// TIA Portal project "Ampelanlage_1" (V20)

(* hardware
DEVICE "S7-1500/ET200MP-Station_1"  S7-1500 station
   slot 0: "Profilschiene_0"  Rack  6ES7 590-1***0-0AA0
   slot 1: "PLC_1"  CPU 1513-1 PN  6ES7 513-1AM03-0AB0  V4.0
      slot 3: "CPU-Display_1"  6ES7591-1AA00-0AA0
      slot 32768: "PROFINET-Schnittstelle_1"  X1
         slot 32769: "Port_1"  X1 P1
         slot 32770: "Port_2"  X1 P2
      slot 34817: "Virtual CP interface port_1"  Virtual CP interface port  Virtual CP interface port FW V4.0
   slot 2: "DI 16x24VDC BA_1"  DI 16x24VDC BA  6ES7 521-1BH10-0AA0  V1.1
   slot 3: "DQ 16x24VDC/0.5A ST_1"  DQ 16x24VDC/0.5A ST  6ES7 522-1BH00-0AB0  V2.0
   slot 4: "AI 8xU/I/R/RTD BA_2"  AI 8xU/I/R/RTD BA  6ES7 531-7QF00-0AB0  V1.0
   slot 5: "AQ 8xU/I HS_2"  AQ 8xU/I HS  6ES7 532-5HF00-0AB0  V2.2
DEVICE "HMI_1"  TP700 Comfort
   slot 0: "HMI_1"  TP700 Comfort  6AV2 124-0GC01-0AX0  17.0.0.0
   slot 1: "HMI_RT_1"  TP700 Comfort  6AV2 124-0GC01-0AX0  17.0.0.0
   slot 5: "HMI_1.IE_CP_1"  PROFINET Interface  17.0.0.0
      slot 1: "PROFINET Schnittstelle_1"  PROFINET Interface
         slot 1: "Port_1"  Port
         slot 2: "Port_2"  Port
   slot 7: "HMI_1.MPI/DP_CP_1"  MPI/DP Interface  17.0.0.0
*)

// ===== PLC "PLC_1"  CPU 1513-1 PN =====

VAR_GLOBAL   // PLC tag table "Eingaenge"
   "S1" AT %E0.0 : Bool;   // Starttaster
END_VAR

VAR_GLOBAL   // PLC tag table "Ausgaenge"
   "1H1" AT %A0.0 : Bool;   // Hauptstraße 1 (rot)
   "1H2" AT %A0.1 : Bool;   // Hauptstraße 1 (gelb)
   "1H3" AT %A0.2 : Bool;   // Hauptstraße 1 (grün)
   "2H1" AT %A0.3 : Bool;   // Hauptstraße 2 (rot)
   "2H2" AT %A0.4 : Bool;   // Hauptstraße 2 (gelb)
   "2H3" AT %A0.5 : Bool;   // Hauptstraße 2 (grün)
   "3H1" AT %A0.6 : Bool;   // Nebenstraße 1 (rot)
   "3H2" AT %A0.7 : Bool;   // Nebenstraße 1 (gelb)
   "3H3" AT %A1.0 : Bool;   // Nebenstraße 1 (grün)
   "4H1" AT %A1.1 : Bool;   // Nebenstraße 2 (rot)
   "4H2" AT %A1.2 : Bool;   // Nebenstraße 2 (gelb)
   "4H3" AT %A1.3 : Bool;   // Nebenstraße 2 (grün)
   "5H1" AT %A1.4 : Bool;   // Fußgänger 1 (rot)
   "5H2" AT %A1.5 : Bool;   // Fußgänger 1 (grün)
   "6H1" AT %A1.6 : Bool;   // Fußgänger 2 (rot)
   "6H2" AT %A1.7 : Bool;   // Fußgänger 2 (grün)
END_VAR

TYPE "typSignale"
   STRUCT
      Hauptstrasse : Struct
         Rot : Bool;   // Hauptstraße Ampel (rot)
         Gelb : Bool;   // Hauptstraße Ampel (gelb)
         Gruen : Bool;   // Hauptstraße Ampel (grün)
      END_STRUCT;
      Nebenstrasse : Struct
         Rot : Bool;   // Nebenstraße Ampel (rot)
         Gelb : Bool;   // Nebenstraße Ampel (gelb)
         Gruen : Bool;   // Nebenstraße Ampel (grün)
      END_STRUCT;
      Fussgaenger : Struct
         Rot : Bool;   // Fußgänger Ampel (rot)
         Gruen : Bool;   // Fußgänger Ampel (grün)
      END_STRUCT;
   END_STRUCT;
END_TYPE

TYPE "typPhasen"
   STRUCT
      Phase_1 : Struct
         NR : UDInt := 1;
         Phasen_Zeit : Time := T#3s;
         Aktiv : Bool;
      END_STRUCT;
      Phase_2 : Struct
         NR : UDInt := 2;
         Phasen_Zeit : Time := T#2s;
         Aktiv : Bool;
      END_STRUCT;
      Phase_3 : Struct
         NR : UDInt := 3;
         Phasen_Zeit : Time := T#10s;
         Aktiv : Bool;
      END_STRUCT;
      Phase_4 : Struct
         NR : UDInt := 4;
         Phasen_Zeit : Time := T#2s;
         Aktiv : Bool;
      END_STRUCT;
      Phase_5 : Struct
         NR : UDInt := 5;
         Phasen_Zeit : Time := T#3s;
         Aktiv : Bool;
      END_STRUCT;
      Phase_6 : Struct
         NR : UDInt := 6;
         Phasen_Zeit : Time := T#2s;
         Aktiv : Bool;
      END_STRUCT;
      Phase_7 : Struct
         NR : UDInt := 7;
         Phasen_Zeit : Time := T#8s;
         Aktiv : Bool;
      END_STRUCT;
      Phase_8 : Struct
         NR : UDInt := 8;
         Phasen_Zeit : Time := T#2s;
         Aktiv : Bool;
      END_STRUCT;
   END_STRUCT;
END_TYPE

TYPE "typTransitionen"
   STRUCT
      Phasen_Transitionen : Struct
         P_1_2 : Bool;
         P_2_3 : Bool;
         P_3_4 : Bool;
         P_4_5 : Bool;
         P_5_6 : Bool;
         P_6_7 : Bool;
         P_7_8 : Bool;
      END_STRUCT;
      Schritt_Transitionen : Struct
         T_0_1 : Bool;
         T_1_2 : Bool;
         T_2_0 : Bool;
         T_2_1 : Bool;
      END_STRUCT;
   END_STRUCT;
END_TYPE

DATA_BLOCK "HMI_Schnittstelle"   // DB1
{ S7_Optimized_Access := 'TRUE' }
VERSION : 0.1
   VAR
      Eingänge : Struct
         S1 : Bool;   // Schalter S1
      END_STRUCT;
      Ausgänge : Struct
         Signale : "typSignale";
      END_STRUCT;
      Schritt_Nr : DInt;
      Ampelphase : Time;
      Phasen : "typPhasen";
      Transitionen : "typTransitionen";
      Anlage_ein : Bool;
   END_VAR
BEGIN
END_DATA_BLOCK

DATA_BLOCK "IDB_Schritte_Ampelanlage"   // DB2
{ S7_Optimized_Access := 'TRUE' }
VERSION : 0.1
// stored: InstanceOfName Prog_Schrittkette_Ampelanlage
"Prog_Schrittkette_Ampelanlage"
BEGIN
END_DATA_BLOCK

FUNCTION_BLOCK "Prog_Schrittkette_Ampelanlage"   // FB1, FBD
{ S7_Optimized_Access := 'TRUE' }
VERSION : 0.1
   VAR_INPUT
      eStart : Bool;
   END_VAR
   VAR_OUTPUT
      aSchritt_Nr : DInt;
   END_VAR
   VAR_IN_OUT
      eaPhasen : "typPhasen";
      eaTransitionen : "typTransitionen";
      eaPhasenzeit : Array[0..8] of Time;
   END_VAR
   VAR
      Schritt_0 : Bool := true;   // 0: Initialschritt
      Schritt_1 : Bool;   // 1: Ampelphase 1
      Schritt_2 : Bool;   // 8: Ampelphase 8
      TOF_Schritt1 : TON_TIME;
      TON_Phase1 : TON_TIME;
      TON_Phase2 : TON_TIME;
      TON_Phase3 : TON_TIME;
      TON_Phase4 : TON_TIME;
      TON_Phase5 : TON_TIME;
      TON_Phase6 : TON_TIME;
      TON_Phase7 : TON_TIME;
      TON_Phase8 : TON_TIME;
      RTRIG_Start_Taster : R_TRIG;
      MDB_Phase_1 : "Ampelphase";
      MDB_Phase_2 : "Ampelphase";
      MDB_Phase_3 : "Ampelphase";
      MDB_Phase_4 : "Ampelphase";
      MDB_Phase_5 : "Ampelphase";
      MDB_Phase_6 : "Ampelphase";
      MDB_Phase_7 : "Ampelphase";
      MDB_Phase_8 : "Ampelphase";
      Phasen_gestartet : Bool;
   END_VAR
BEGIN

REGION Network 1: Anlage in Grundstellung
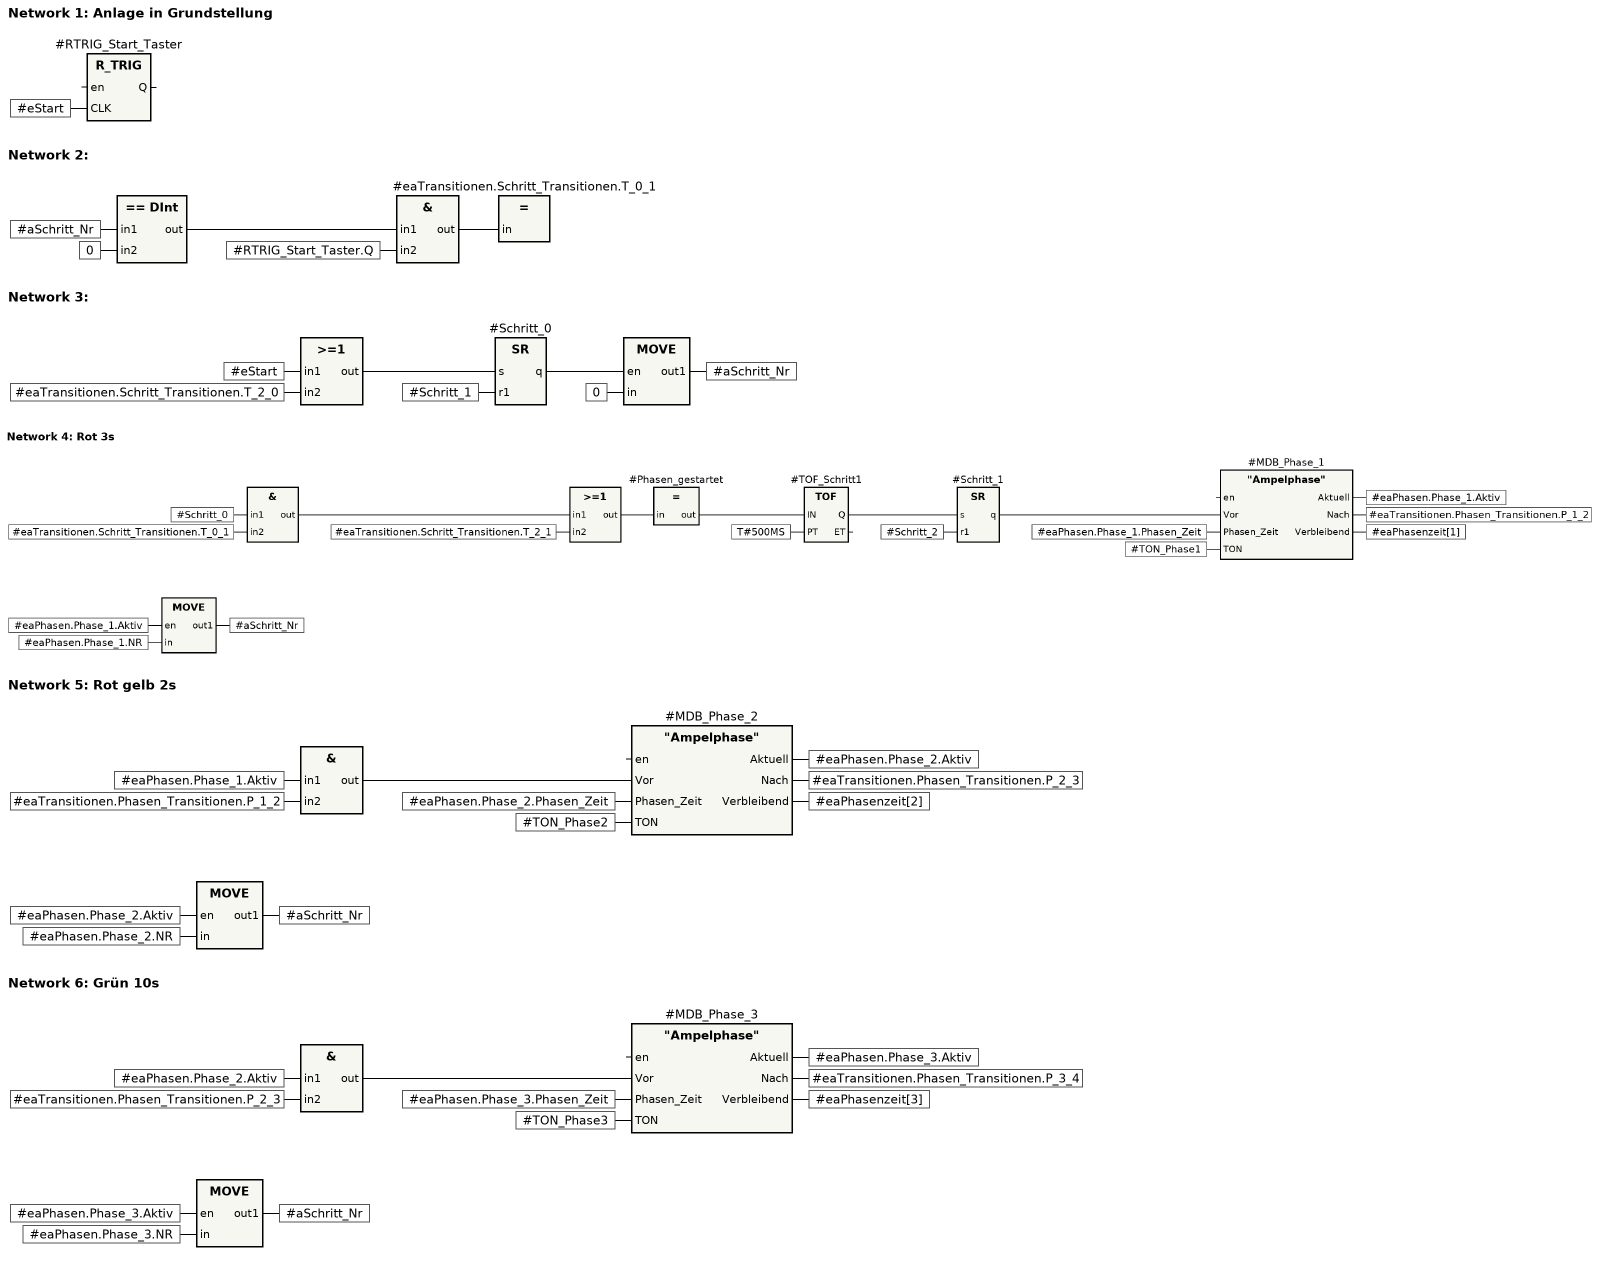
   #RTRIG_Start_Taster(CLK := #eStart);   // R_TRIG
END_REGION

REGION Network 2
   #eaTransitionen.Schritt_Transitionen.T_0_1 := (#aSchritt_Nr = 0) AND #RTRIG_Start_Taster.Q;
END_REGION

REGION Network 3
   IF #eStart OR #eaTransitionen.Schritt_Transitionen.T_2_0 THEN
       #Schritt_0 := TRUE;   // SR flip-flop
   END_IF;
   IF #Schritt_1 THEN #Schritt_0 := FALSE; END_IF;
   IF #Schritt_0 THEN #aSchritt_Nr := 0; END_IF;
END_REGION

REGION Network 4: Rot 3s
   #Phasen_gestartet := (#Schritt_0 AND #eaTransitionen.Schritt_Transitionen.T_0_1) OR #eaTransitionen.Schritt_Transitionen.T_2_1;
   #TOF_Schritt1(IN := #Phasen_gestartet, PT := T#500MS);   // TOF
   IF #TOF_Schritt1.Q THEN
       #Schritt_1 := TRUE;   // SR flip-flop
   END_IF;
   IF #Schritt_2 THEN #Schritt_1 := FALSE; END_IF;
   #MDB_Phase_1(Vor := #Schritt_1,   // "Ampelphase"
                Phasen_Zeit := #eaPhasen.Phase_1.Phasen_Zeit,
                TON := #TON_Phase1,
                Aktuell => #eaPhasen.Phase_1.Aktiv,
                Nach => #eaTransitionen.Phasen_Transitionen.P_1_2,
                Verbleibend => #eaPhasenzeit[1]);
   IF #eaPhasen.Phase_1.Aktiv THEN #aSchritt_Nr := #eaPhasen.Phase_1.NR; END_IF;
END_REGION

REGION Network 5: Rot gelb 2s
   #MDB_Phase_2(Vor := #eaPhasen.Phase_1.Aktiv AND #eaTransitionen.Phasen_Transitionen.P_1_2,   // "Ampelphase"
                Phasen_Zeit := #eaPhasen.Phase_2.Phasen_Zeit,
                TON := #TON_Phase2,
                Aktuell => #eaPhasen.Phase_2.Aktiv,
                Nach => #eaTransitionen.Phasen_Transitionen.P_2_3,
                Verbleibend => #eaPhasenzeit[2]);
   IF #eaPhasen.Phase_2.Aktiv THEN #aSchritt_Nr := #eaPhasen.Phase_2.NR; END_IF;
END_REGION

REGION Network 6: Grün 10s
   #MDB_Phase_3(Vor := #eaPhasen.Phase_2.Aktiv AND #eaTransitionen.Phasen_Transitionen.P_2_3,   // "Ampelphase"
                Phasen_Zeit := #eaPhasen.Phase_3.Phasen_Zeit,
                TON := #TON_Phase3,
                Aktuell => #eaPhasen.Phase_3.Aktiv,
                Nach => #eaTransitionen.Phasen_Transitionen.P_3_4,
                Verbleibend => #eaPhasenzeit[3]);
   IF #eaPhasen.Phase_3.Aktiv THEN #aSchritt_Nr := #eaPhasen.Phase_3.NR; END_IF;
END_REGION

REGION Network 7: Gelb 2s
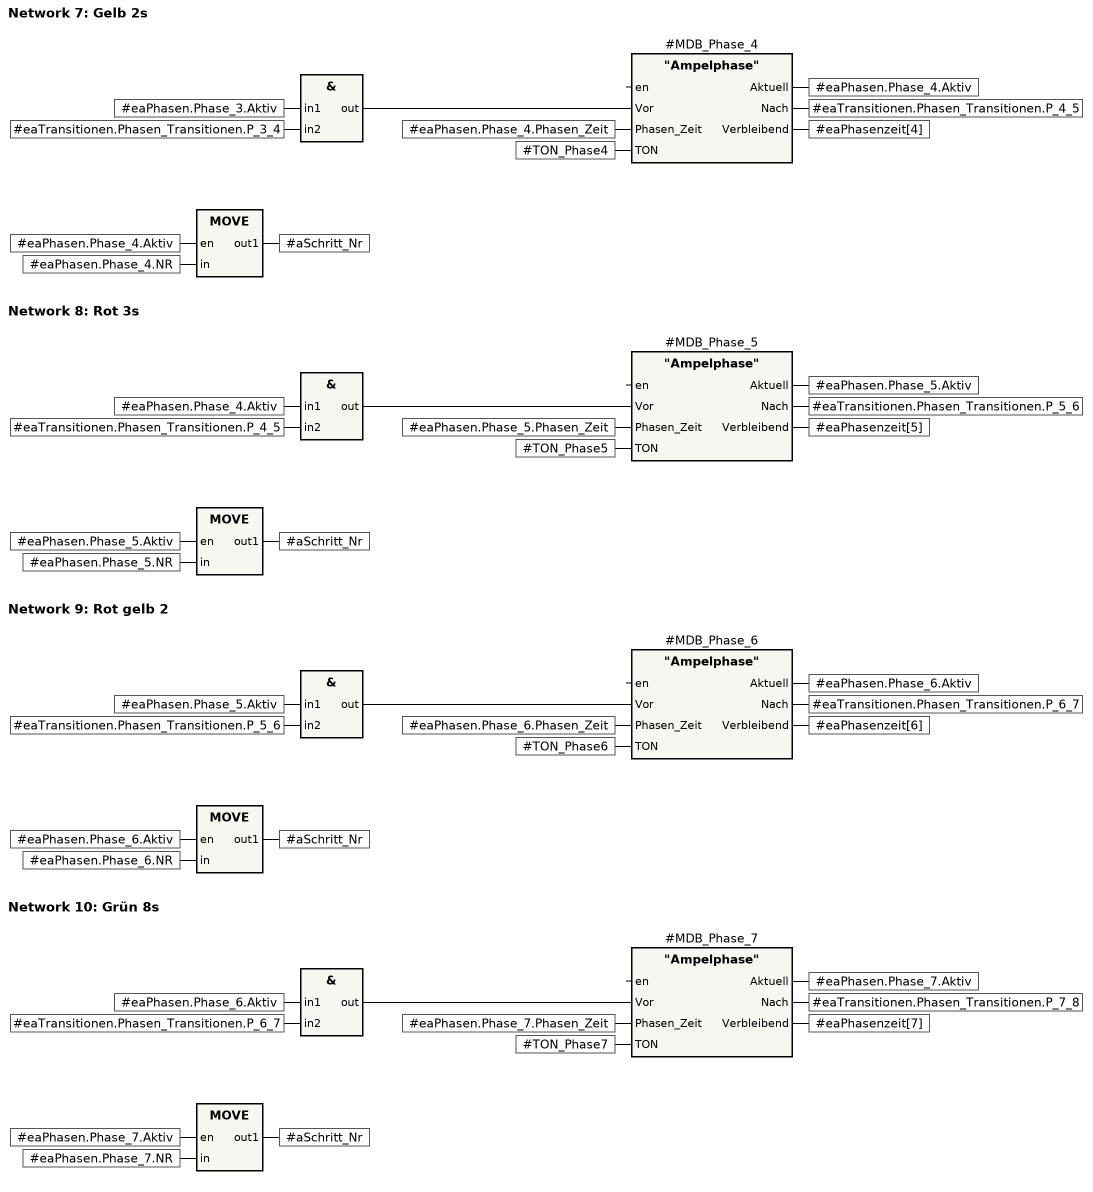
   #MDB_Phase_4(Vor := #eaPhasen.Phase_3.Aktiv AND #eaTransitionen.Phasen_Transitionen.P_3_4,   // "Ampelphase"
                Phasen_Zeit := #eaPhasen.Phase_4.Phasen_Zeit,
                TON := #TON_Phase4,
                Aktuell => #eaPhasen.Phase_4.Aktiv,
                Nach => #eaTransitionen.Phasen_Transitionen.P_4_5,
                Verbleibend => #eaPhasenzeit[4]);
   IF #eaPhasen.Phase_4.Aktiv THEN #aSchritt_Nr := #eaPhasen.Phase_4.NR; END_IF;
END_REGION

REGION Network 8: Rot 3s
   #MDB_Phase_5(Vor := #eaPhasen.Phase_4.Aktiv AND #eaTransitionen.Phasen_Transitionen.P_4_5,   // "Ampelphase"
                Phasen_Zeit := #eaPhasen.Phase_5.Phasen_Zeit,
                TON := #TON_Phase5,
                Aktuell => #eaPhasen.Phase_5.Aktiv,
                Nach => #eaTransitionen.Phasen_Transitionen.P_5_6,
                Verbleibend => #eaPhasenzeit[5]);
   IF #eaPhasen.Phase_5.Aktiv THEN #aSchritt_Nr := #eaPhasen.Phase_5.NR; END_IF;
END_REGION

REGION Network 9: Rot gelb 2
   #MDB_Phase_6(Vor := #eaPhasen.Phase_5.Aktiv AND #eaTransitionen.Phasen_Transitionen.P_5_6,   // "Ampelphase"
                Phasen_Zeit := #eaPhasen.Phase_6.Phasen_Zeit,
                TON := #TON_Phase6,
                Aktuell => #eaPhasen.Phase_6.Aktiv,
                Nach => #eaTransitionen.Phasen_Transitionen.P_6_7,
                Verbleibend => #eaPhasenzeit[6]);
   IF #eaPhasen.Phase_6.Aktiv THEN #aSchritt_Nr := #eaPhasen.Phase_6.NR; END_IF;
END_REGION

REGION Network 10: Grün 8s
   #MDB_Phase_7(Vor := #eaPhasen.Phase_6.Aktiv AND #eaTransitionen.Phasen_Transitionen.P_6_7,   // "Ampelphase"
                Phasen_Zeit := #eaPhasen.Phase_7.Phasen_Zeit,
                TON := #TON_Phase7,
                Aktuell => #eaPhasen.Phase_7.Aktiv,
                Nach => #eaTransitionen.Phasen_Transitionen.P_7_8,
                Verbleibend => #eaPhasenzeit[7]);
   IF #eaPhasen.Phase_7.Aktiv THEN #aSchritt_Nr := #eaPhasen.Phase_7.NR; END_IF;
END_REGION

REGION Network 11: Gelb 2s
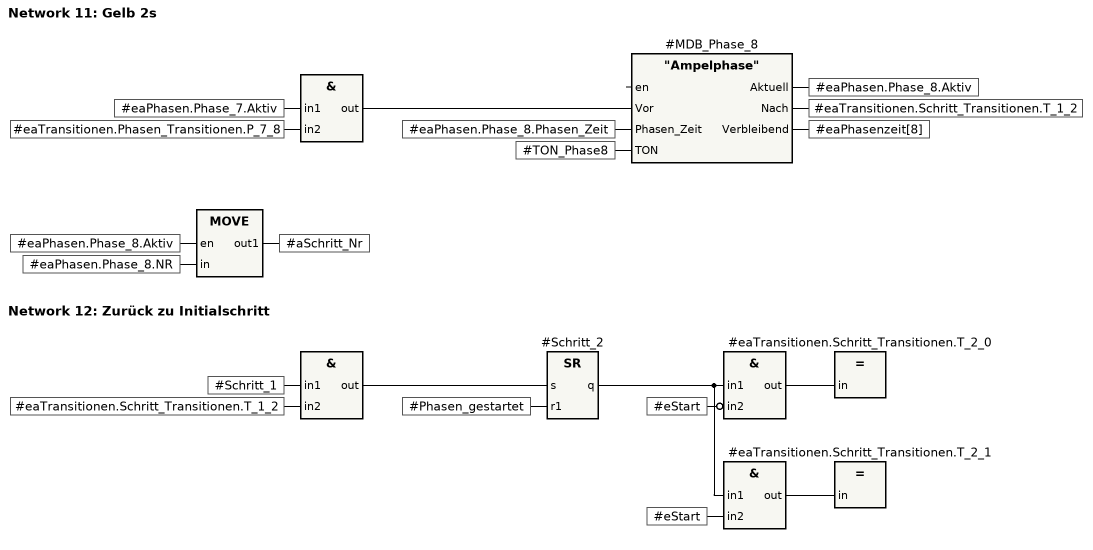
   #MDB_Phase_8(Vor := #eaPhasen.Phase_7.Aktiv AND #eaTransitionen.Phasen_Transitionen.P_7_8,   // "Ampelphase"
                Phasen_Zeit := #eaPhasen.Phase_8.Phasen_Zeit,
                TON := #TON_Phase8,
                Aktuell => #eaPhasen.Phase_8.Aktiv,
                Nach => #eaTransitionen.Schritt_Transitionen.T_1_2,
                Verbleibend => #eaPhasenzeit[8]);
   IF #eaPhasen.Phase_8.Aktiv THEN #aSchritt_Nr := #eaPhasen.Phase_8.NR; END_IF;
END_REGION

REGION Network 12: Zurück zu Initialschritt
   IF #Schritt_1 AND #eaTransitionen.Schritt_Transitionen.T_1_2 THEN
       #Schritt_2 := TRUE;   // SR flip-flop
   END_IF;
   IF #Phasen_gestartet THEN #Schritt_2 := FALSE; END_IF;
   #eaTransitionen.Schritt_Transitionen.T_2_0 := #Schritt_2 AND NOT #eStart;
   #eaTransitionen.Schritt_Transitionen.T_2_1 := #Schritt_2 AND #eStart;
END_REGION
END_FUNCTION_BLOCK

FUNCTION_BLOCK "Ampelphase"   // FB2, FBD
{ S7_Optimized_Access := 'TRUE' }
VERSION : 0.1
   VAR_INPUT
      Vor : Bool;
      Phasen_Zeit : Time;
   END_VAR
   VAR_OUTPUT
      Aktuell : Bool;
      Nach : Bool;
      Verbleibend : Time;
   END_VAR
   VAR_IN_OUT
      TON : TON_TIME;
   END_VAR
BEGIN

REGION Network 1
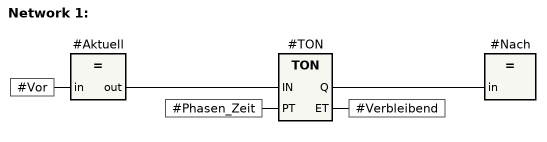
   #Aktuell := #Vor;
   #TON(IN := #Vor, PT := #Phasen_Zeit, ET => #Verbleibend);   // TON
   #Nach := #TON.Q;
END_REGION
END_FUNCTION_BLOCK

FUNCTION_BLOCK "Anlagensignale_einlesen"   // FB3, FBD
{ S7_Optimized_Access := 'TRUE' }
VERSION : 0.1
   VAR
      RTRIG_HMI_Taster : R_TRIG;
      RTRIG_eStart : R_TRIG;
   END_VAR
BEGIN

REGION Network 1: Flankenabfragen
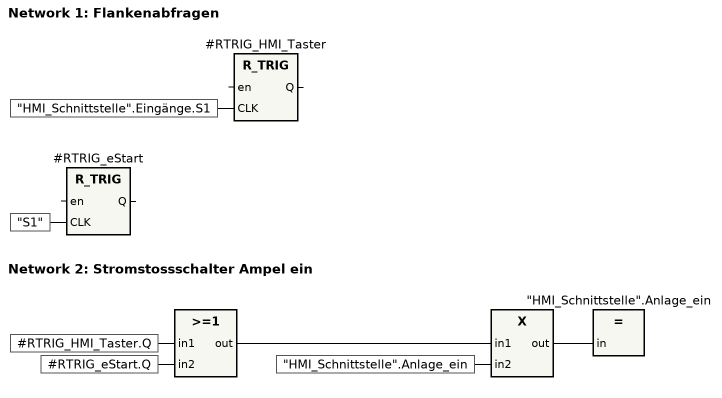
   #RTRIG_HMI_Taster(CLK := "HMI_Schnittstelle".Eingänge.S1);   // R_TRIG
   #RTRIG_eStart(CLK := "S1");   // R_TRIG
END_REGION

REGION Network 2: Stromstossschalter Ampel ein
   "HMI_Schnittstelle".Anlage_ein := (#RTRIG_HMI_Taster.Q OR #RTRIG_eStart.Q) XOR "HMI_Schnittstelle".Anlage_ein;
END_REGION
END_FUNCTION_BLOCK

FUNCTION_BLOCK "Takt"   // FB10101, FBD
TITLE = Taktbaustein parametrierbar
{ S7_Optimized_Access := 'TRUE' }
VERSION : 0.1
// ACHTUNG: keine Zeit darf 0ms sein, ansonsten funktioniert der Baustein nicht.
   VAR_INPUT
      ePulsZeit : Time := T#500MS;   // So lange ist Ausgang = TRUE
      ePauseZeit : Time := T#500MS;   // So lange ist Ausgang = FALSE
   END_VAR
   VAR_OUTPUT
      Q : Bool;
   END_VAR
   VAR
      TP_Puls : TP_TIME;
      TP_Pause : TP_TIME;
   END_VAR
BEGIN

REGION Network 1: Puls Timer
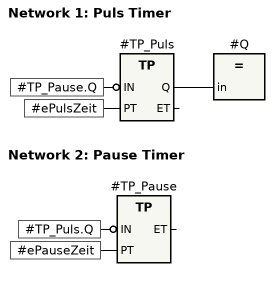
   #TP_Puls(IN := NOT #TP_Pause.Q, PT := #ePulsZeit);   // TP
   #Q := #TP_Puls.Q;
END_REGION

REGION Network 2: Pause Timer
   #TP_Pause(IN := NOT #TP_Puls.Q, PT := #ePauseZeit);   // TP
END_REGION
END_FUNCTION_BLOCK

FUNCTION "Aus_an_Anlage" : Void   // FC1, FBD
{ S7_Optimized_Access := 'TRUE' }
VERSION : 0.1
   VAR_INPUT
      eSignale : "typSignale";
   END_VAR
BEGIN

REGION Network 1: Ampeln Hauptstraße
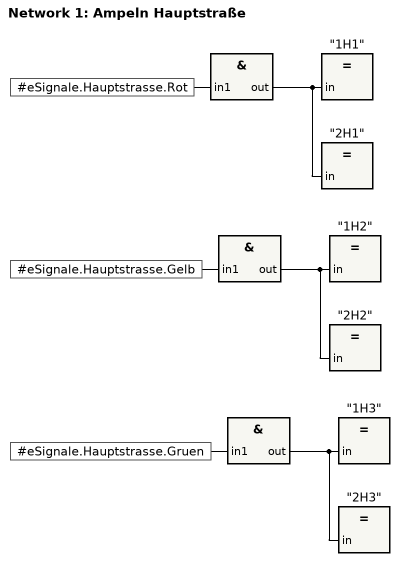
   "1H1" := #eSignale.Hauptstrasse.Rot;
   "2H1" := #eSignale.Hauptstrasse.Rot;
   "1H2" := #eSignale.Hauptstrasse.Gelb;
   "2H2" := #eSignale.Hauptstrasse.Gelb;
   "1H3" := #eSignale.Hauptstrasse.Gruen;
   "2H3" := #eSignale.Hauptstrasse.Gruen;
END_REGION

REGION Network 2 (SCL): Nebenstraße 1 (rot)
   // Ampel Nebenstraße

   "3H1" := "4H1" := #eSignale.Nebenstrasse.Rot;
   "3H2" := "4H2" := #eSignale.Nebenstrasse.Gelb;
   "3H3" := "4H3" := #eSignale.Nebenstrasse.Gruen;


   // Ampel Fussgaenger
   "5H1" := "6H1" := #eSignale.Fussgaenger.Rot;
   "5H2" := "6H2" := #eSignale.Fussgaenger.Gruen;
END_REGION
END_FUNCTION

FUNCTION "Aus_Ampelanlage" : Void   // FC2, FBD
{ S7_Optimized_Access := 'TRUE' }
VERSION : 0.1
   VAR_INPUT
      eSchritt_Nr : DInt;
   END_VAR
   VAR_OUTPUT
      aSignale : "typSignale";
   END_VAR
   VAR_TEMP
      Initialschritt : Bool;
   END_VAR
BEGIN

REGION Network 1
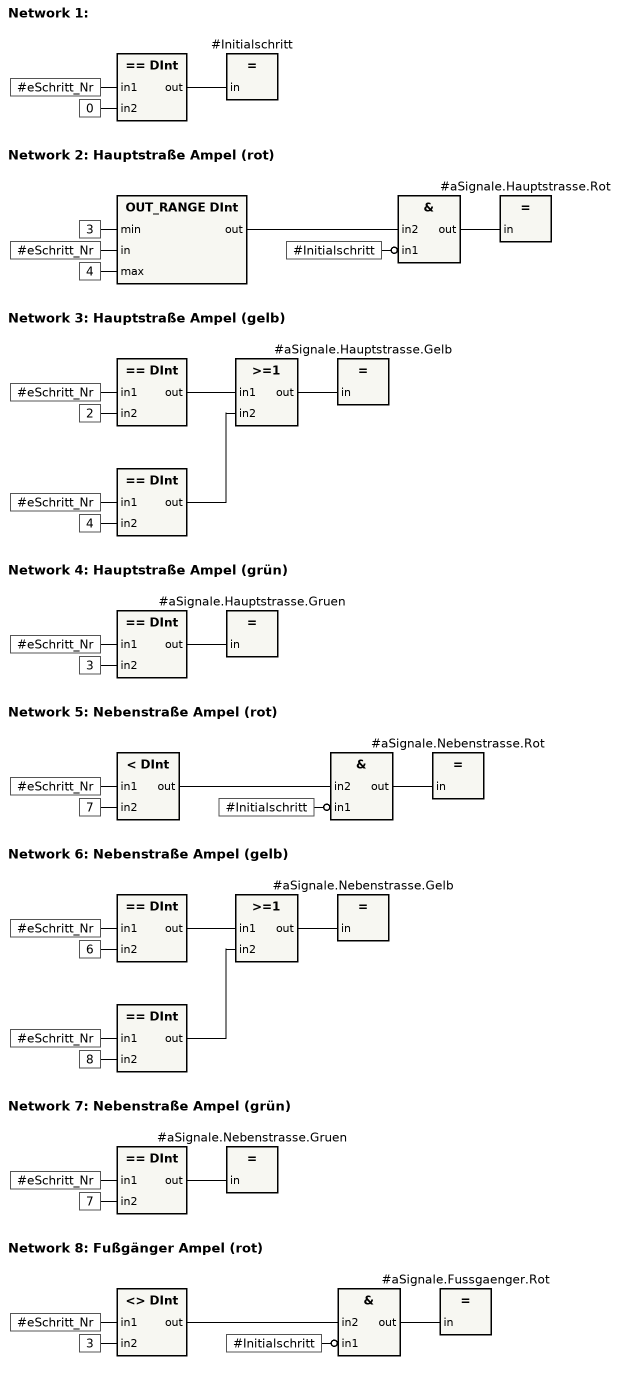
   #Initialschritt := #eSchritt_Nr = 0;
END_REGION

REGION Network 2: Hauptstraße Ampel (rot)
   #aSignale.Hauptstrasse.Rot := ((#eSchritt_Nr < 3) OR (#eSchritt_Nr > 4)) AND NOT #Initialschritt;
END_REGION

REGION Network 3: Hauptstraße Ampel (gelb)
   #aSignale.Hauptstrasse.Gelb := (#eSchritt_Nr = 2) OR (#eSchritt_Nr = 4);
END_REGION

REGION Network 4: Hauptstraße Ampel (grün)
   #aSignale.Hauptstrasse.Gruen := #eSchritt_Nr = 3;
END_REGION

REGION Network 5: Nebenstraße Ampel (rot)
   #aSignale.Nebenstrasse.Rot := (#eSchritt_Nr < 7) AND NOT #Initialschritt;
END_REGION

REGION Network 6: Nebenstraße Ampel (gelb)
   #aSignale.Nebenstrasse.Gelb := (#eSchritt_Nr = 6) OR (#eSchritt_Nr = 8);
END_REGION

REGION Network 7: Nebenstraße Ampel (grün)
   #aSignale.Nebenstrasse.Gruen := #eSchritt_Nr = 7;
END_REGION

REGION Network 8: Fußgänger Ampel (rot)
   #aSignale.Fussgaenger.Rot := (#eSchritt_Nr <> 3) AND NOT #Initialschritt;
END_REGION

REGION Network 9: Fußgänger Ampel (grün)
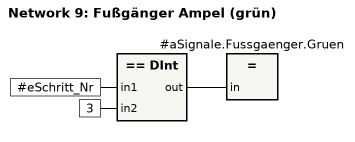
   #aSignale.Fussgaenger.Gruen := #eSchritt_Nr = 3;
END_REGION
END_FUNCTION

ORGANIZATION_BLOCK "Main"   // OB1, FBD, ProgramCycle
TITLE = "Main Program Sweep (Cycle)"
{ S7_Optimized_Access := 'TRUE' }
VERSION : 0.1
   VAR_INPUT
      Initial_Call : Bool;   // Initial call of this OB
      Remanence : Bool;   // =True, if remanent data are available
   END_VAR
   VAR_TEMP
      Phasenzeit : Array[0..8] of Time;
   END_VAR
BEGIN

REGION Network 1
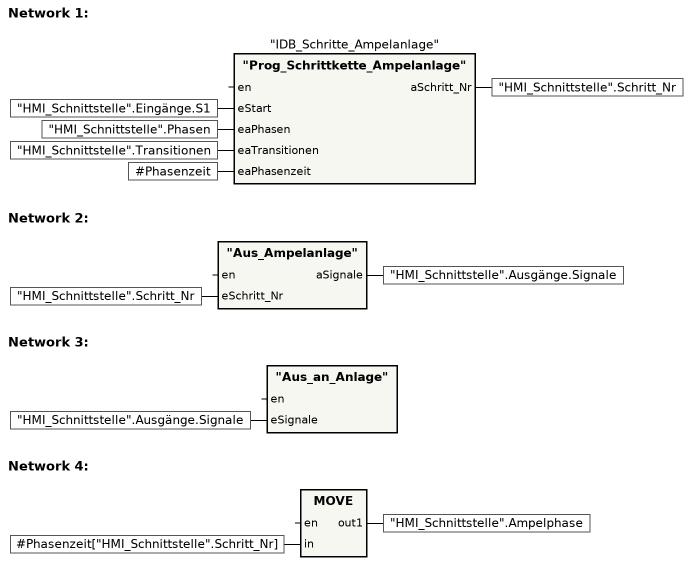
   "IDB_Schritte_Ampelanlage"(eStart := "HMI_Schnittstelle".Eingänge.S1,   // "Prog_Schrittkette_Ampelanlage"
                           eaPhasen := "HMI_Schnittstelle".Phasen,
                           eaTransitionen := "HMI_Schnittstelle".Transitionen,
                           eaPhasenzeit := #Phasenzeit,
                           aSchritt_Nr => "HMI_Schnittstelle".Schritt_Nr);
END_REGION

REGION Network 2
   "Aus_Ampelanlage"(eSchritt_Nr := "HMI_Schnittstelle".Schritt_Nr,
                     aSignale => "HMI_Schnittstelle".Ausgänge.Signale);
END_REGION

REGION Network 3
   "Aus_an_Anlage"(eSignale := "HMI_Schnittstelle".Ausgänge.Signale);
END_REGION

REGION Network 4
   "HMI_Schnittstelle".Ampelphase := #Phasenzeit["HMI_Schnittstelle".Schritt_Nr];
END_REGION
END_ORGANIZATION_BLOCK

(* ===== HMI "HMI_RT_1" =====
system functions are stored by id; their names below are inferred from use
connection "HMI_Verbindung_1": ETHERNET, S7_1500_OMS

HMI tags "Standard-Variablentabelle"
   "HMI_Schnittstelle_S1" : Bool = PLC HMI_Schnittstelle.Eingänge.S1, 500 ms
   "HMI_Schnittstelle_Ausgänge_Schritt_Nr" : DInt = PLC HMI_Schnittstelle.Schritt_Nr, 100 ms
   "HMI_Schnittstelle_Ausgänge_1H1" : Bool = PLC HMI_Schnittstelle.Ausgänge.Signale.Hauptstrasse.Rot, 100 ms
   "HMI_Schnittstelle_Ausgänge_1H2" : Bool = PLC HMI_Schnittstelle.Ausgänge.Signale.Hauptstrasse.Gelb, 100 ms
   "HMI_Schnittstelle_Ausgänge_1H3" : Bool = PLC HMI_Schnittstelle.Ausgänge.Signale.Hauptstrasse.Gruen, 100 ms
   "HMI_Schnittstelle_Ausgänge_2H1" : Bool = PLC HMI_Schnittstelle.Ausgänge.Signale.Nebenstrasse.Rot, 100 ms
   "HMI_Schnittstelle_Ausgänge_2H2" : Bool = PLC HMI_Schnittstelle.Ausgänge.Signale.Nebenstrasse.Gelb, 100 ms
   "HMI_Schnittstelle_Ausgänge_2H3" : Bool = PLC HMI_Schnittstelle.Ausgänge.Signale.Nebenstrasse.Gruen, 100 ms
   "HMI_Schnittstelle_Ausgänge_3H1" : Bool = PLC HMI_Schnittstelle.Ausgänge.Signale.Fussgaenger.Rot, 100 ms
   "HMI_Schnittstelle_Ausgänge_3H2" : Bool = PLC HMI_Schnittstelle.Ausgänge.Signale.Fussgaenger.Gruen, 100 ms
   "HMI_Schnittstelle_Ampelphase" : Time = PLC HMI_Schnittstelle.Ampelphase, 100 ms

screen "Ampelanlage" 800x480
   Button "Schaltfläche_1" at 700,444 size 96x32; TextOff 'S1'
      on Click: InvertBit("HMI_Schnittstelle_S1")
      Appearance <- "HMI_Schnittstelle_S1"
   Circle "Kreis_1" at 286,238 size 16x16
      Appearance <- "HMI_Schnittstelle_Ausgänge_1H1"
   Circle "Kreis_2" at 268,238 size 16x16
      Appearance <- "HMI_Schnittstelle_Ausgänge_1H2"
   Circle "Kreis_3" at 250,238 size 16x16
      Appearance <- "HMI_Schnittstelle_Ausgänge_1H3"
   Circle "Kreis_4" at 498,26 size 16x16
      Appearance <- "HMI_Schnittstelle_Ausgänge_1H1"
   Circle "Kreis_5" at 516,26 size 16x16
      Appearance <- "HMI_Schnittstelle_Ausgänge_1H2"
   Circle "Kreis_6" at 534,26 size 16x16
      Appearance <- "HMI_Schnittstelle_Ausgänge_1H3"
   Circle "Kreis_7" at 498,318 size 16x16
      Appearance <- "HMI_Schnittstelle_Ausgänge_2H1"
   Circle "Kreis_8" at 498,336 size 16x16
      Appearance <- "HMI_Schnittstelle_Ausgänge_2H2"
   Circle "Kreis_9" at 498,354 size 16x16
      Appearance <- "HMI_Schnittstelle_Ausgänge_2H3"
   Circle "Kreis_10" at 286,298 size 16x16
      Appearance <- "HMI_Schnittstelle_Ausgänge_3H1"
   Circle "Kreis_11" at 268,298 size 16x16
      Appearance <- "HMI_Schnittstelle_Ausgänge_3H2"
   Circle "Kreis_12" at 516,238 size 16x16
      Appearance <- "HMI_Schnittstelle_Ausgänge_3H2"
   Circle "Kreis_13" at 498,238 size 16x16
      Appearance <- "HMI_Schnittstelle_Ausgänge_3H1"
   IOField "EA-Feld_1" at 4,444 size 96x32; FormatPattern 9
      ProcessValue <- "HMI_Schnittstelle_Ausgänge_Schritt_Nr"
   TextField "Textfeld_1" at 4,420 size 101x23; Text 'Schritt-Nr.'
   IOField "EA-Feld_2" at 352,144 size 96x32; FormatPattern 99999; Unit  ms
      ProcessValue <- "HMI_Schnittstelle_Ampelphase"
   TextField "Textfeld_2" at 347,120 size 105x23; Text 'Phasenzeit'
*)